   IOField "I/O field_37" at 183,323 size 90x29; Authorization "Commissioning"; FormatPattern 999; Unit  step
      ProcessValue <- "2110_BTCS_CNTRL_DB_BTCS_STEP"
   Button "HmiScreenItemData_10" at 43,323 size 137x29; TextOn 'Back'; TextOff 'BWTS Step'
   Button "HmiScreenItemData_51" at 43,358 size 137x29; TextOn 'Back'; TextOff 'BWTS State'
   Button "HmiScreenItemData_54" at 276,323 size 532x29; TextOn 'Back'; TextOff 'IGG STEP'; TextList "STEP LIST BTCS"
      ProcessValue <- "2110_BTCS_CNTRL_DB_BTCS_STEP"
   Button "HmiScreenItemData_55" at 276,358 size 532x29; TextOn 'Back'; TextOff 'IGG STEP'; TextList "STATE LIST BTCS"
      ProcessValue <- "2110_BTCS_CNTRL_DB_BTCS_STATE"
   Circle "Circle_2" at 421,496 size 26x26
      Appearance <- "80_From_HMI_BWT_BYPASS"
   Button "HmiScreenItemData_57" at 88,494 size 304x33; TextOn 'Back'; TextOff 'Ballast Water Treatment'; Authorization "Operate"
      on Press: InvertBit("80_From_HMI_BWT_BYPASS(1)"); ResetBit("80_From_HMI_CRG_BLNK_MODE(1)")
      Appearance <- "80_From_HMI_BWT_BYPASS(1)"
      ObjectEnable <- "100_GCU_AUTO_SEQ_DB_CRNT_STEP"
   Circle "Circle_3" at 421,534 size 26x26
      Appearance <- "80_From_HMI_CRG_BLNK_MODE"
   Button "HmiScreenItemData_58" at 88,532 size 304x33; TextOn 'Back'; TextOff 'Cargo Blanketing'; Authorization "Operate"
      on Press: InvertBit("80_From_HMI_CRG_BLNK_MODE(1)"); ResetBit("80_From_HMI_BWT_BYPASS(1)")
      Appearance <- "80_From_HMI_CRG_BLNK_MODE(1)"
      ObjectEnable <- "100_GCU_AUTO_SEQ_DB_CRNT_STEP"
   Button "HmiScreenItemData_56" at 41,461 size 425x27; TextOn 'Back'; TextOff 'Inert Gas Transfer Mode'
   Button "Button_7" at 817,526 size 79x32; TextOff '1'; Authorization "Operate"
      Appearance <- "504_Tank Grouping_DB2020_GROUP ACTIVE INT 1"
      on Press: function_b14e0dd5("504_Tank Grouping_DB2020_GROUP ACTIV 1", 0)
   Button "Button_8" at 817,560 size 79x32; TextOff '2'; Authorization "Operate"
      Appearance <- "504_Tank Grouping_DB2020_GROUP ACTIVE INT 2"
      on Press: function_b14e0dd5("504_Tank Grouping_DB2020_GROUP ACTIV 2", 0)
   Button "Button_9" at 493,539 size 100x23; TextOff 'TANK - 1P'; Authorization "Operate"
      on Press: function_b14e0dd5("504_Tank Grouping_DB2020_TANK ACTIV 2", 0)
      Appearance <- "504_Tank Grouping_DB2020_TANK ACTIV 2"
   Button "Button_14" at 493,571 size 100x23; TextOff 'TANK - 2P'; Authorization "Operate"
      on Press: function_b14e0dd5("504_Tank Grouping_DB2020_TANK ACTIV 4", 0)
      Appearance <- "504_Tank Grouping_DB2020_TANK ACTIV 4"
   Button "Button_15" at 493,603 size 100x23; TextOff 'TANK - 3P'; Authorization "Operate"
      on Press: function_b14e0dd5("504_Tank Grouping_DB2020_TANK ACTIV 6", 0)
      Appearance <- "504_Tank Grouping_DB2020_TANK ACTIV 6"
   Button "Button_16" at 493,636 size 100x23; TextOff 'TANK - 4P'; Authorization "Operate"
      on Press: function_b14e0dd5("504_Tank Grouping_DB2020_TANK ACTIV 8", 0)
      Appearance <- "504_Tank Grouping_DB2020_TANK ACTIV 8"
   Button "Button_17" at 493,668 size 100x23; TextOff 'TANK - 5P'; Authorization "Operate"
      on Press: function_b14e0dd5("504_Tank Grouping_DB2020_TANK ACTIV 10", 0)
      Appearance <- "504_Tank Grouping_DB2020_TANK ACTIV 10"
   Button "Button_18" at 493,700 size 100x23; TextOff 'TANK - 6P'; Authorization "Operate"
      on Press: function_b14e0dd5("504_Tank Grouping_DB2020_TANK ACTIV 12", 0)
      Appearance <- "504_Tank Grouping_DB2020_TANK ACTIV 12"
   Button "Button_19" at 493,733 size 100x23; TextOff 'TANK - APT'; Authorization "Operate"
      on Press: function_b14e0dd5("504_Tank Grouping_DB2020_TANK ACTIV 14", 0)
      Appearance <- "504_Tank Grouping_DB2020_TANK ACTIV 14"
   Button "Button_20" at 706,539 size 100x23; TextOff 'TANK - 1S'; Authorization "Operate"
      on Press: function_b14e0dd5("504_Tank Grouping_DB2020_TANK ACTIV 3", 0)
      Appearance <- "504_Tank Grouping_DB2020_TANK ACTIV 3"
   Button "Button_21" at 706,571 size 100x23; TextOff 'TANK - 2S'; Authorization "Operate"
      on Press: function_b14e0dd5("504_Tank Grouping_DB2020_TANK ACTIV 5", 0)
      Appearance <- "504_Tank Grouping_DB2020_TANK ACTIV 5"
   Button "Button_22" at 706,603 size 100x23; TextOff 'TANK - 3S'; Authorization "Operate"
      on Press: function_b14e0dd5("504_Tank Grouping_DB2020_TANK ACTIV 7", 0)
      Appearance <- "504_Tank Grouping_DB2020_TANK ACTIV 7"
   Button "Button_23" at 706,635 size 100x23; TextOff 'TANK - 4S'; Authorization "Operate"
      on Press: function_b14e0dd5("504_Tank Grouping_DB2020_TANK ACTIV 9", 0)
      Appearance <- "504_Tank Grouping_DB2020_TANK ACTIV 9"
   Button "Button_24" at 706,667 size 100x23; TextOff 'TANK - 5S'; Authorization "Operate"
      on Press: function_b14e0dd5("504_Tank Grouping_DB2020_TANK ACTIV 11", 0)
      Appearance <- "504_Tank Grouping_DB2020_TANK ACTIV 11"
   Button "Button_25" at 706,700 size 100x23; TextOff 'TANK - 6S'; Authorization "Operate"
      on Press: function_b14e0dd5("504_Tank Grouping_DB2020_TANK ACTIV 13", 0)
      Appearance <- "504_Tank Grouping_DB2020_TANK ACTIV 13"
   IOField "I/O field_38" at 183,358 size 90x29; Authorization "Commissioning"; FormatPattern 9; Unit  state
      ProcessValue <- "2110_BTCS_CNTRL_DB_BTCS_STATE"
   Switch "Switch_8" at 776,732 size 32x29; CaptionText 'Switch'; TextOn 'ON'; TextOff 'OFF'; Authorization "User administration"; PictureOff "Design_5_PilotLight_Green_Off"; PictureOn "Design_5_PilotLight_Green_On"
      on Change: InvertBit("80_From_HMI_Test Tank Request")
      ProcessValue <- "504_Tank Grouping_DB2020_RUN"
   Circle "Circle_31" at 621,507 size 20x20
      Appearance <- "504_Tank Grouping_DB2020_RUN TANK 1"
      Visibility <- "504_Tank Grouping_DB2020_RUN TANK 1"
   Circle "Circle_4" at 600,573 size 20x20
      Appearance <- "504_Tank Grouping_DB2020_GROUP of TANK 4"
   Circle "Circle_6" at 599,604 size 20x20
      Appearance <- "504_Tank Grouping_DB2020_GROUP of TANK 6"
   Circle "Circle_7" at 599,541 size 20x20
      Appearance <- "504_Tank Grouping_DB2020_GROUP of TANK 2"
   Circle "Circle_8" at 599,669 size 20x20
      Appearance <- "504_Tank Grouping_DB2020_GROUP of TANK 10"
   Circle "Circle_10" at 599,637 size 20x20
      Appearance <- "504_Tank Grouping_DB2020_GROUP of TANK 8"
   Circle "Circle_11" at 599,734 size 20x20
      Appearance <- "504_Tank Grouping_DB2020_GROUP of TANK 14"
   Circle "Circle_12" at 599,701 size 20x20
      Appearance <- "504_Tank Grouping_DB2020_GROUP of TANK 12"
   IOField "I/O field_8" at 599,544 size 20x14; FormatPattern 99
      ProcessValue <- "504_Tank Grouping_DB2020_GROUP of TANK 2"
   IOField "I/O field_9" at 599,576 size 20x14; FormatPattern 99
      ProcessValue <- "504_Tank Grouping_DB2020_GROUP of TANK 4"
   IOField "I/O field_26" at 599,607 size 20x14; FormatPattern 99
      ProcessValue <- "504_Tank Grouping_DB2020_GROUP of TANK 6"
   IOField "I/O field_28" at 599,640 size 20x14; FormatPattern 99
      ProcessValue <- "504_Tank Grouping_DB2020_GROUP of TANK 8"
   IOField "I/O field_30" at 599,672 size 20x14; FormatPattern 99
      ProcessValue <- "504_Tank Grouping_DB2020_GROUP of TANK 10"
   IOField "I/O field_33" at 599,704 size 20x14; FormatPattern 99
      ProcessValue <- "504_Tank Grouping_DB2020_GROUP of TANK 12"
   IOField "I/O field_35" at 599,737 size 20x14; FormatPattern 99
      ProcessValue <- "504_Tank Grouping_DB2020_GROUP of TANK 14"
   Circle "Circle_13" at 678,573 size 20x20
      Appearance <- "504_Tank Grouping_DB2020_GROUP of TANK 5"
   Circle "Circle_14" at 678,603 size 20x20
      Appearance <- "504_Tank Grouping_DB2020_GROUP of TANK 7"
   Circle "Circle_15" at 678,541 size 20x20
      Appearance <- "504_Tank Grouping_DB2020_GROUP of TANK 3"
   Circle "Circle_16" at 678,668 size 20x20
      Appearance <- "504_Tank Grouping_DB2020_GROUP of TANK 11"
   Circle "Circle_17" at 678,636 size 20x20
      Appearance <- "504_Tank Grouping_DB2020_GROUP of TANK 9"
   Circle "Circle_18" at 678,701 size 20x20
      Appearance <- "504_Tank Grouping_DB2020_GROUP of TANK 13"
   IOField "I/O field_23" at 678,544 size 20x14; FormatPattern 99
      ProcessValue <- "504_Tank Grouping_DB2020_GROUP of TANK 3"
   IOField "I/O field_24" at 678,576 size 20x14; FormatPattern 99
      ProcessValue <- "504_Tank Grouping_DB2020_GROUP of TANK 5"
   IOField "I/O field_27" at 678,606 size 20x14; FormatPattern 99
      ProcessValue <- "504_Tank Grouping_DB2020_GROUP of TANK 7"
   IOField "I/O field_29" at 678,639 size 20x14; FormatPattern 99
      ProcessValue <- "504_Tank Grouping_DB2020_GROUP of TANK 9"
   IOField "I/O field_32" at 678,671 size 20x14; FormatPattern 99
      ProcessValue <- "504_Tank Grouping_DB2020_GROUP of TANK 11"
   IOField "I/O field_34" at 678,704 size 20x14; FormatPattern 99
      ProcessValue <- "504_Tank Grouping_DB2020_GROUP of TANK 13"
   Circle "Circle_32" at 621,540 size 20x20
      Appearance <- "504_Tank Grouping_DB2020_RUN TANK 2"
      Visibility <- "504_Tank Grouping_DB2020_RUN TANK 2"
   Circle "Circle_33" at 656,540 size 20x20
      Appearance <- "504_Tank Grouping_DB2020_RUN TANK 3"
      Visibility <- "504_Tank Grouping_DB2020_RUN TANK 3"
   Circle "Circle_34" at 621,572 size 20x20
      Appearance <- "504_Tank Grouping_DB2020_RUN TANK 4"
      Visibility <- "504_Tank Grouping_DB2020_RUN TANK 4"
   Circle "Circle_35" at 656,572 size 20x20
      Appearance <- "504_Tank Grouping_DB2020_RUN TANK 5"
      Visibility <- "504_Tank Grouping_DB2020_RUN TANK 5"
   Circle "Circle_36" at 621,604 size 20x20
      Appearance <- "504_Tank Grouping_DB2020_RUN TANK 6"
      Visibility <- "504_Tank Grouping_DB2020_RUN TANK 6"
   Circle "Circle_37" at 656,604 size 20x20
      Appearance <- "504_Tank Grouping_DB2020_RUN TANK 7"
      Visibility <- "504_Tank Grouping_DB2020_RUN TANK 7"
   Circle "Circle_38" at 621,636 size 20x20
      Appearance <- "504_Tank Grouping_DB2020_RUN TANK 8"
      Visibility <- "504_Tank Grouping_DB2020_RUN TANK 8"
   Circle "Circle_39" at 656,636 size 20x20
      Appearance <- "504_Tank Grouping_DB2020_RUN TANK 9"
      Visibility <- "504_Tank Grouping_DB2020_RUN TANK 9"
   Circle "Circle_40" at 621,668 size 20x20
      Appearance <- "504_Tank Grouping_DB2020_RUN TANK 10"
      Visibility <- "504_Tank Grouping_DB2020_RUN TANK 10"
   Circle "Circle_41" at 656,668 size 20x20
      Appearance <- "504_Tank Grouping_DB2020_RUN TANK 11"
      Visibility <- "504_Tank Grouping_DB2020_RUN TANK 11"
   Circle "Circle_42" at 621,701 size 20x20
      Appearance <- "504_Tank Grouping_DB2020_RUN TANK 12"
      Visibility <- "504_Tank Grouping_DB2020_RUN TANK 12"
   Circle "Circle_43" at 656,701 size 20x20
      Appearance <- "504_Tank Grouping_DB2020_RUN TANK 13"
      Visibility <- "504_Tank Grouping_DB2020_RUN TANK 13"
   Circle "Circle_44" at 621,733 size 20x20
      Appearance <- "504_Tank Grouping_DB2020_RUN TANK 14"
      Visibility <- "504_Tank Grouping_DB2020_RUN TANK 14"
   TextField "Text field_7" at 648,740 size 136x18; Text 'Test Tank Request'
   Rectangle "Rectangle_6" at 816,488 size 82x37
      Visibility <- "504_Tank Grouping_DB2020_SetGroupSR"
   Button "Button_13" at 819,491 size 76x31; TextOff 'Set Group'; Authorization "Parameter Change"
      Appearance <- "504_Tank Grouping_DB2020_GROUP SET"
      on Press: function_b14e0dd5("504_Tank Grouping_DB2020_SetGroup", 0)
   Button "HmiScreenItemData_5" at 41,576 size 426x27; TextOn 'Back'; TextOff 'Automatic Gas to Tank Valves Cycling'
   Button "HmiScreenItemData_19" at 371,722 size 83x35; TextOn 'ENABLE'; TextOff 'Enable'; Authorization "Operating Mode"
      on Press: InvertBit("504_Tank Grouping_DB2020_Valve Cycle_Enable")
      Appearance <- "504_Tank Grouping_DB2020_Valve Cycle_Enable"
   TextField "Text field_8" at 54,652 size 254x18; Text 'Gas to Tank Valves Cycle Frequency'
   TextField "Text field_9" at 54,690 size 233x18; Text 'Gas to Tank Valves Cycle Length'
   TextField "Text field_10" at 54,618 size 85x18; Text 'Description'
   TextField "Text field_12" at 311,618 size 67x18; Text 'Setpoint'
   IOField "I/O field_39" at 310,649 size 70x28; Authorization "Operate"; FormatPattern 999; Unit h
      ProcessValue <- "504_Tank Grouping_DB2020_Valve Cycle_Period"
   IOField "I/O field_40" at 310,685 size 70x28; Authorization "Operate"; FormatPattern 9999; Unit s
      ProcessValue <- "504_Tank Grouping_DB2020_Valve Cycle_Length"
   TextField "Text field_13" at 385,618 size 58x18; Text 'Elapsed'
   IOField "I/O field_41" at 384,649 size 70x28; Authorization "Operate"; FormatPattern 999; Unit h
      ProcessValue <- "504_Tank Grouping_DB2020_Cycle Period_ET"
   IOField "I/O field_42" at 384,685 size 70x28; Authorization "Operate"; FormatPattern 9999; Unit s
      ProcessValue <- "504_Tank Grouping_DB2020_Cycle Length_ET"
   IOField "I/O field_48" at 1172,169 size 33x28; Authorization "User administration"; FormatPattern 99; Unit h
      ProcessValue <- "Sequence Times_DB_Treatment Timer_Hours Left"
   IOField "I/O field_51" at 1140,169 size 33x28; Authorization "User administration"; FormatPattern 99; Unit d
      ProcessValue <- "Sequence Times_DB_Treatment Timer_Days Left"
   IOField "I/O field_52" at 1204,169 size 35x28; Authorization "User administration"; FormatPattern 99; Unit m
      ProcessValue <- "Sequence Times_DB_Treatment Timer_Minutes Left"
   IOField "I/O field_43" at 1156,201 size 83x28; Authorization "User administration"; FormatPattern 999; Unit  min
      ProcessValue <- "504_Tank Grouping_DB2020_Diff Time Remain"
      Visibility <- "AlwaysTRUE"
   IOField "I/O field_44" at 1204,233 size 35x28; Authorization "User administration"; FormatPattern 99; Unit m
      ProcessValue <- "Sequence Times_DB_Pre-Dwell Timer_Minutes Left"
   IOField "I/O field_45" at 1172,233 size 33x28; Authorization "User administration"; FormatPattern 99; Unit h
      ProcessValue <- "Sequence Times_DB_Pre-Dwell Timer_Hours Left"
   IOField "I/O field_46" at 1140,233 size 33x28; Authorization "User administration"; FormatPattern 99; Unit d
      ProcessValue <- "Sequence Times_DB_Pre-Dwell Timer_Days Left"
   IOField "I/O field_47" at 1040,132 size 92x28; Authorization "Operating Mode"; FormatPattern 999.9; Unit  Days
      ProcessValue <- "Sequence Times_DB_Jurney Time"
   IOField "I/O field_49" at 1072,169 size 33x28; Authorization "User administration"; FormatPattern 99; Unit h
      ProcessValue <- "Sequence Times_DB_Treatment Timer_Hours"
   IOField "I/O field_50" at 1040,169 size 33x28; Authorization "User administration"; FormatPattern 99; Unit d
      ProcessValue <- "Sequence Times_DB_Treatment Timer_Days"
   IOField "I/O field_53" at 1104,169 size 35x28; Authorization "User administration"; FormatPattern 99; Unit m
      ProcessValue <- "Sequence Times_DB_Treatment Timer_Minutes"
   IOField "I/O field_54" at 1172,132 size 33x28; Authorization "User administration"; FormatPattern 99; Unit h
      ProcessValue <- "Sequence Times_DB_Jurney Timer_Hours Left"
   IOField "I/O field_55" at 1133,132 size 40x28; Authorization "User administration"; FormatPattern 999; Unit d
      ProcessValue <- "Sequence Times_DB_Jurney Timer_Days Left"
   IOField "I/O field_56" at 1204,132 size 35x28; Authorization "User administration"; FormatPattern 99; Unit m
      ProcessValue <- "Sequence Times_DB_Jurney Timer_Minutes Left"
   IOField "I/O field_57" at 1040,233 size 79x28; Authorization "Commissioning"; FormatPattern 9999.9; Unit  Hrs
      ProcessValue <- "Sequence Times_DB_Pre-Dwell Time"
   IOField "I/O field_58" at 1040,267 size 79x28; Authorization "Commissioning"; FormatPattern 999.9; Unit  Hrs
      ProcessValue <- "Sequence Times_DB_De-Ox Time"
   IOField "I/O field_59" at 1204,267 size 35x28; Authorization "User administration"; FormatPattern 99; Unit m
      ProcessValue <- "Sequence Times_DB_De-Ox Timer_Minutes Left"
   IOField "I/O field_60" at 1172,267 size 33x28; Authorization "User administration"; FormatPattern 99; Unit h
      ProcessValue <- "Sequence Times_DB_De-Ox Timer_Hours Left"
   IOField "I/O field_61" at 1140,267 size 33x28; Authorization "User administration"; FormatPattern 99; Unit d
      ProcessValue <- "Sequence Times_DB_De-Ox Timer_Days Left"
   IOField "I/O field_62" at 1040,301 size 79x28; Authorization "Commissioning"; FormatPattern 999.9; Unit  Hrs
      ProcessValue <- "Sequence Times_DB_De-Ox SP Time"
   IOField "I/O field_63" at 1040,335 size 79x28; Authorization "Commissioning"; FormatPattern 999.9; Unit  Hrs
      ProcessValue <- "Sequence Times_DB_Dwell Time"
   IOField "I/O field_64" at 1204,335 size 35x28; Authorization "User administration"; FormatPattern 99; Unit m
      ProcessValue <- "Sequence Times_DB_Dwell Timer_Minutes Left"
   IOField "I/O field_65" at 1172,335 size 33x28; Authorization "User administration"; FormatPattern 99; Unit h
      ProcessValue <- "Sequence Times_DB_Dwell Timer_Hours Left"
   IOField "I/O field_66" at 1140,335 size 33x28; Authorization "User administration"; FormatPattern 99; Unit d
      ProcessValue <- "Sequence Times_DB_Dwell Timer_Days Left"
   IOField "I/O field_2" at 1040,369 size 79x28; Authorization "Commissioning"; FormatPattern 999.9; Unit  Hrs
      ProcessValue <- "Sequence Times_DB_Re-Ox Time"
   IOField "I/O field_67" at 1204,369 size 35x28; Authorization "User administration"; FormatPattern 99; Unit m
      ProcessValue <- "Sequence Times_DB_Re-Ox Timer_Minutes Left"
   IOField "I/O field_68" at 1172,369 size 33x28; Authorization "User administration"; FormatPattern 99; Unit h
      ProcessValue <- "Sequence Times_DB_Re-Ox Timer_Hours Left"
   IOField "I/O field_69" at 1140,369 size 33x28; Authorization "User administration"; FormatPattern 99; Unit d
      ProcessValue <- "Sequence Times_DB_Re-Ox Timer_Days Left"
   IOField "I/O field_70" at 1040,403 size 79x28; Authorization "Commissioning"; FormatPattern 999.9; Unit  Hrs
      ProcessValue <- "Sequence Times_DB_Post-Dwell Time"
   IOField "I/O field_71" at 1204,403 size 35x28; Authorization "User administration"; FormatPattern 99; Unit m
      ProcessValue <- "Sequence Times_DB_Post-Dwell Timer_Minutes Left"
   IOField "I/O field_72" at 1172,403 size 33x28; Authorization "User administration"; FormatPattern 99; Unit h
      ProcessValue <- "Sequence Times_DB_Post-Dwell Timer_Hours Left"
   IOField "I/O field_73" at 1140,403 size 33x28; Authorization "User administration"; FormatPattern 99; Unit d
      ProcessValue <- "Sequence Times_DB_Post-Dwell Timer_Days Left"
   TextField "Text field_15" at 621,419 size 156x18; Text 'Treatment Timer Test'
      Visibility <- "user_group"
   Circle "Circle_5" at 599,507 size 20x20
      Appearance <- "504_Tank Grouping_DB2020_GROUP of TANK 1"
   IOField "I/O field_7" at 599,510 size 20x14; FormatPattern 99
      ProcessValue <- "504_Tank Grouping_DB2020_GROUP of TANK 1"
   Button "HmiScreenItemData_50" at 1156,297 size 83x35; TextOn 'Back'; TextOff 'Boost'; Authorization "Commissioning"
      on Press: InvertBit("Sequence Times_DB_Boost")
      Visibility <- "user_group"
      Appearance <- "Sequence Times_DB_Boost"
   TextField "Text field_16" at 38,419 size 76x18; Text 'HeartBeat'
      Visibility <- "user_group"
   TextField "Text field_18" at 201,422 size 107x18; Text 'PLC HeartBeat'
      Visibility <- "user_group"
   Circle "Circle_45" at 6,412 size 26x26
      Appearance <- "IGG HMI HEART BEAT"
   Circle "Circle_46" at 166,414 size 26x26
      Appearance <- "IGG PLC HEART BEAT"
   Switch "Switch_1" at 774,411 size 32x29; CaptionText 'Switch'; TextOn 'ON'; TextOff 'OFF'; Authorization "User administration"; PictureOff "Design_5_PilotLight_Green_Off"; PictureOn "Design_5_PilotLight_Green_On"
      on Change: InvertBit("80_From_HMI_Jurney Start Simulator")
      Visibility <- "user_group"
      ProcessValue <- "80_From_HMI_Jurney Start Simulator"
   TextField "Text field_19" at 445,403 size 133x18; Text 'Log IGG Simulator'
      Visibility <- "user_group"
   Switch "Switch_2" at 568,393 size 32x29; CaptionText 'Switch'; TextOn 'ON'; TextOff 'OFF'; Authorization "User administration"; PictureOff "Design_5_PilotLight_Green_Off"; PictureOn "Design_5_PilotLight_Green_On"
      on Change: InvertBit("68_Sys_Status_Data_LOG IGG Simulator")
      Visibility <- "user_group"
      ProcessValue <- "68_Sys_Status_Data_LOG IGG Simulator"
   TextField "Text field_20" at 445,435 size 136x18; Text 'Log GCU Simulator'
      Visibility <- "user_group"
   Switch "Switch_3" at 568,425 size 32x29; CaptionText 'Switch'; TextOn 'ON'; TextOff 'OFF'; Authorization "User administration"; PictureOff "Design_5_PilotLight_Green_Off"; PictureOn "Design_5_PilotLight_Green_On"
      on Change: InvertBit("68_Sys_Status_Data_LOG GCU Simulator")
      Visibility <- "user_group"
      ProcessValue <- "68_Sys_Status_Data_LOG GCU Simulator"
   Button "Button_5" at 53,722 size 210x35; TextOff 'PGC Setpoint Protection'
      on Press: function_efd93a16("PGC Setpoint Protection", 400, 200, -1, -1, 1)
   Button "Button_26" at 280,114 size 209x107; TextOff 'Text'
      on Release: function_efd93a16("Salinity - Acceptance", 168, 315, -1, 0, 1)
      Visibility <- "2068_Sys_Status_Data_SAL_VALID"
   Button "Button_27" at 283,115 size 204x107; TextOff 'Text'
      on Release: function_efd93a16("Tank Times", 300, 200, -1, 0, 1)
      Visibility <- "2068_Sys_Status_Data_Times Visibil"
   Group "Group_1" at 909,732 size 329x37
   IOField "I/O field_74" at 1172,201 size 33x28; Authorization "User administration"; FormatPattern 99; Unit h
      ProcessValue <- "Sequence Times_DB_Offset Timer_Hours Left"
   IOField "I/O field_75" at 1140,201 size 33x28; Authorization "User administration"; FormatPattern 99; Unit d
      ProcessValue <- "Sequence Times_DB_Offset Timer_Days Left"
   IOField "I/O field_76" at 1204,201 size 35x28; Authorization "User administration"; FormatPattern 99; Unit m
      ProcessValue <- "Sequence Times_DB_Offset Timer_Minutes Left"
   Circle "Circle_23" at 762,90 size 24x24
      Appearance <- "2110_BTCS_CNTRL_DB_BTCS_STEP"
   Circle "Circle_24" at 762,119 size 24x24
      Appearance <- "100_GCU_AUTO_SEQ_DB_CRNT_STEP"
   Circle "Circle_25" at 762,149 size 24x24
      Appearance <- "2110_BTCS_CNTRL_DB_BTCS_STEP"
   Circle "Circle_26" at 762,179 size 24x24
      Appearance <- "2110_BTCS_CNTRL_DB_BTCS_STEP"
   Circle "Circle_27" at 762,209 size 24x24
      Appearance <- "100_GCU_AUTO_SEQ_DB_CRNT_STEP"
   Circle "Circle_28" at 762,239 size 24x24
      Appearance <- "2110_BTCS_CNTRL_DB_BTCS_STEP"
   Circle "Circle_29" at 762,269 size 24x24
      Appearance <- "2110_BTCS_CNTRL_DB_BTCS_STEP"
   TextField "Text field_34" at 980,733 size 187x35; Text 'TIMES VALID'
      Visibility <- "2102_TIME_CALCS_DB_TIMES_VALID"
   TextField "Text field_4" at 909,732 size 329x37; Text 'TIMES INVALID'
      Visibility <- "2102_TIME_CALCS_DB_TIMES_VALID"
   Rectangle "Rectangle_27" at 921,659 size 322x40
      Visibility <- "2068_Sys_Status_Data_SAL_CNF_CHK"
   TextField "Text field_62" at 925,664 size 156x30; Text 'Confirm Salinity? :'
      Visibility <- "2068_Sys_Status_Data_SAL_CNF_CHK"
   Button "Button_6" at 1086,664 size 67x30; TextOff 'YES'
      on Press: function_b14e0dd5("80_From_HMI_LOW_SAL_ACPT", 0)
      Visibility <- "2068_Sys_Status_Data_SAL_CNF_CHK"
   Button "Button_3" at 1166,664 size 67x30; TextOff 'NO'
      on Press: function_b14e0dd5("80_From_HMI_LOW_SAL_RJCT", 0)
      Visibility <- "2068_Sys_Status_Data_SAL_CNF_CHK"
   Rectangle "Rectangle_28" at 916,659 size 327x40
      Visibility <- "2100_AUTO_SEQ_DB_SEQ_RNG"
      Appearance <- "2102_TIME_CALCS_DB_RE_OX_SP_TMR_DN"
   TextField "Text field_49" at 920,664 size 211x30; Text 'Salinity Value :'
      Visibility <- "2100_AUTO_SEQ_DB_SEQ_RNG"
   IOField "I/O field_36" at 1131,664 size 95x30; Authorization "Operate"; FormatPattern 99.9; Unit psu
      Visibility <- "2100_AUTO_SEQ_DB_SEQ_RNG"
      ProcessValue <- "80_From_HMI_SAL_VALUE"

PopupScreen "SD Card overflow" 665x230
   Button "Button_1" at 0,0 size 665x230; TextOff 'Data Logging SD Card Memory Full'
      on Click: function_efd93a16("SD Card overflow", 0, 0, -1, -1, 1)
      on Press: ResetBit("Logging SD Card Overflow")

PopupScreen "Salinity - Fresh Water Alert" 1280x800
   Button "Button_1" at 115,225 size 1050x284; TextOff 'NOTE: BALLAST WATER SALINITY IS FRESH WATER LEVEL This System Is Not Certified For FRESH WATER Treatment. Do Wish To Continue Ballast Water Treatment?'
   Button "Button_2" at 666,514 size 105x50; TextOff 'NO'
      on Release: ActivateScreen("Balast Water Treatment Setup", 0)
      on Press: function_b14e0dd5("80_From_HMI_LOW_SAL_RJCT", 0)
   Button "Button_3" at 500,514 size 105x50; TextOff 'YES'
      on Release: ActivateScreen("Balast Water Treatment Setup", 0)
      on Press: function_b14e0dd5("80_From_HMI_LOW_SAL_ACPT", 0)

screen "Main Page" 1280x800, template "Template"
   GraphicView "Graphic view_49" at 158,415 size 30x45; Picture "Graphic_72"
   GraphicView "Graphic view_20" at 140,368 size 380x356; Picture "IGG_6"
   GraphicView "Graphic view_62" at 134,449 size 92x8; Picture "Graphic_20"
   GraphicView "Graphic view_5" at 464,423 size 90x19; Picture "Graphic_82"
   GraphicView "Graphic view_41" at 228,459 size 9x40; Picture "Graphic_57"
   GraphicView "Graphic view_40" at 222,449 size 15x13; Picture "Graphic_41"
   GraphicView "Graphic view_21" at 210,503 size 17x7; Picture "Graphic_63"
   GraphicView "Graphic view_22" at 207,499 size 8x9; Picture "Graphic_64"
   GraphicView "Graphic view_23" at 206,399 size 6x104; Picture "Graphic_70"
   GraphicView "Graphic view_39" at 138,535 size 6x7; Picture "Graphic_70"
   GraphicView "Graphic view_38" at 139,539 size 7x9; Picture "Graphic_64"
   GraphicView "Graphic view_18" at 204,397 size 9x10; Picture "Graphic_67"
   Group "Group_3" at 158,415 size 30x41; Picture "Graphic_72"
   GraphicView "Graphic view_65" at 144,542 size 8x6; Picture "Graphic_63"
   GraphicView "Graphic view_69" at 295,453 size 14x15; Picture "Graphic_36"
   GraphicView "Graphic view_70" at 335,462 size 14x15; Picture "Graphic_36"
   GraphicView "Graphic view_71" at 251,443 size 14x17; Picture "Graphic_79"
   GraphicView "Graphic view_36" at 517,373 size 35x50; Picture "Graphic_108"
   GraphicView "Graphic view_4" at 333,376 size 31x49; Picture "Graphic_108"
   GraphicView "Graphic view_72" at 387,407 size 14x17; Picture "Graphic_36"
   GraphicView "Graphic view_37" at 136,525 size 8x11; Picture "Graphic_67"
   GraphicView "Graphic view_89" at 440,407 size 14x17; Picture "Graphic_36"
   Line "Line_4" at 226,517 size 2x15
      Visibility <- "14_DQ_Data_X001ControlOut"
   GraphicView "Graphic view_84" at 215,511 size 27x55; Picture "Graphic_129"
      Visibility <- "102_Pilot_Burner_DB_FLM_DET"
   GraphicView "Graphic view_90" at 488,409 size 14x15; Picture "Graphic_36"
   GraphicView "Graphic view_1" at 342,415 size 18x41; Picture "Graphic_17"
   GraphicView "Graphic view_60" at 526,412 size 18x41; Picture "Graphic_17"
   GraphicView "Graphic view_82" at 210,499 size 167x147; Picture "Graphic_130"
      Visibility <- "103_Main_Burner_DB_DN_OK(1)"
   IOField "I/O field_17" at 231,558 size 46x17; FormatPattern 999; Unit %
      Visibility <- "10 DI_DATA_FD001_OK"
      ProcessValue <- "12_AI_Data_FD001FlameSignalIn"
   GraphicView "Graphic view_63" at 133,396 size 75x7; Picture "Graphic_63"
   GraphicView "Graphic view_25" at 659,340 size 25x46; Picture "Graphic_148"
   Group "Group_10" at 659,340 size 26x47; Picture "Graphic_148"
   Group "Group_11" at 649,372 size 56x37; Picture "Graphic_224"
   GraphicView "Graphic view_26" at 649,373 size 55x36; Picture "Graphic_224"
   GraphicView "Graphic view_27" at 569,502 size 205x15; Picture "Graphic_232"
   GraphicView "Graphic view_3" at 78,471 size 64x14; Picture "Graphic_82"
   GraphicView "Graphic view_19" at 776,616 size 64x10; Picture "Graphic_82"
   GraphicIOField "Graphic I/O field_2" at 0,485 size 128x131; PictureList "IA Compressor_1"
      ProcessValue <- "82_To_HMI_CA Blower Animation"
   GraphicView "Graphic view_7" at 700,602 size 119x212; Picture "Graphic_150"
   Group "Group" at 133,368 size 421x356; Picture "Graphic_20"
   GraphicView "Graphic view_2" at 821,493 size 449x266; Picture "Graphic_185"
   GraphicView "Graphic view_6" at 68,470 size 18x21; Picture "Graphic_66"
   GraphicView "Graphic view_8" at 41,328 size 96x93; Picture "Graphic_246"
   GraphicView "Graphic view_14" at 630,544 size 17x40; Picture "Graphic_271"
   GraphicView "Graphic view_15" at 570,390 size 205x15; Picture "Graphic_232"
   GraphicView "Graphic view_16" at 561,391 size 26x27; Picture "Graphic_178"
   GraphicView "Graphic view_17" at 757,380 size 17x35; Picture "Graphic_280"
   GraphicView "Graphic view_9" at 525,539 size 156x153; Picture "Graphic_251"
   GraphicView "Graphic view_24" at 561,407 size 14x167; Picture "Graphic_231"
   GraphicView "Graphic view_11" at 555,635 size 21x22; Picture "Graphic_265"
   GraphicView "Graphic view_12" at 555,653 size 29x31; Picture "Graphic_266"
   GraphicView "Graphic view_13" at 572,667 size 133x18; Picture "Graphic_232"
   GraphicView "Graphic view_10" at 549,422 size 26x38; Picture "Graphic_169"
   Group "Group_12" at 649,340 size 56x69; Picture "Graphic_148"
   GraphicView "Graphic view_28" at 756,492 size 17x35; Picture "Graphic_280"
   Group "Group_4" at 648,452 size 56x69; Picture "Graphic_148"
   GraphicView "Graphic view_29" at 658,452 size 25x46; Picture "Graphic_148"
   Group "Group_1" at 658,452 size 26x47; Picture "Graphic_148"
   Group "Group_2" at 648,484 size 56x37; Picture "Graphic_224"
   GraphicView "Graphic view_30" at 648,485 size 55x36; Picture "Graphic_224"

screen "GCU Analogue Inputs" 1280x800, template "Template"
   on GenerateScreen: "TitleUpdater"()
   Button "HmiScreenItemData_1" at 1,1 size 150x43; TextOn 'Back'; TextOff 'Commissioning'
      on Release: ActivateScreen("Commissioning Main Page", 0)
   TextField "Text field_6" at 7,150 size 53x22; Text 'IW800'
   TextField "Text field_8" at 7,270 size 53x22; Text 'IW806'
   TextField "Text field_10" at 7,310 size 53x22; Text 'IW808'
   TextField "Text field_12" at 7,430 size 53x22; Text 'IW814'
   TextField "Text field_30" at 1203,124 size 74x20; Text 'High High'
   TextField "Text field_54" at 649,719 size 228x62; Text 'Note: CSW = Cooling Sea Water'
   TextField "Text field_32" at 7,231 size 53x22; Text 'IW804'
   TextField "Text field_34" at 7,391 size 53x22; Text 'IW812'
   TextField "Text field_36" at 8,191 size 53x22; Text 'IW802'
   TextField "Text field_38" at 8,349 size 53x22; Text 'IW810'
   AlarmView "Alarm view_1" at 0,777 size 1280x23
   IOField "I/O field_62" at 1208,191 size 60x22; FormatPattern 9.9
      ProcessValue <- "84_Setpoints_E400_PT002_HighHigh"
   IOField "I/O field_61" at 1140,191 size 60x22; FormatPattern 9.9
      ProcessValue <- "84_Setpoints_E400_PT002_High"
   TextField "Text field_82" at 60,150 size 220x22; Text 'LIT304 GCU LEVEL'
   TextField "Text field_90" at 286,124 size 64x20; Text 'Reading'
   IOField "I/O field_2" at 287,150 size 70x22; FormatPattern 999; Unit  %
      ProcessValue <- "12_AI_Data_LIT_304_SCALED"
   TextField "Text field_1" at 359,124 size 68x20; Text 'Low Low'
   IOField "I/O field_1" at 361,150 size 60x22; Authorization "Parameter Change"; FormatPattern 999
      ProcessValue <- "19_AUTO_CMNDS_Data_LIT304_CMND_LowLow"
   TextField "Text field_2" at 442,124 size 37x20; Text 'Low'
   IOField "I/O field_3" at 429,150 size 60x22; Authorization "Parameter Change"; FormatPattern 999
      ProcessValue <- "19_AUTO_CMNDS_Data_LIT304_CMND_Low"
   TextField "Text field_3" at 509,124 size 37x20; Text 'High'
   IOField "I/O field_4" at 497,150 size 60x22; Authorization "Parameter Change"; FormatPattern 999
      ProcessValue <- "19_AUTO_CMNDS_Data_LIT304_CMND_High"
   TextField "Text field_4" at 561,124 size 74x20; Text 'High High'
   IOField "I/O field_5" at 565,150 size 60x22; Authorization "Parameter Change"; FormatPattern 999
      ProcessValue <- "19_AUTO_CMNDS_Data_LIT304_CMND_HighHigh"
   TextField "Text field_5" at 434,100 size 76x20; Text 'Setpoints'
   TextField "Text field_7" at 60,270 size 220x22; Text 'TIT406 GAS TO DECK TEMP'
   IOField "I/O field_6" at 287,270 size 70x22; FormatPattern s999; Unit  °C
      ProcessValue <- "12_AI_Data_TIT_406_SCALED"
   IOField "I/O field_7" at 361,270 size 60x22; FormatPattern 999
   IOField "I/O field_8" at 429,270 size 60x22; FormatPattern 999
   IOField "I/O field_9" at 497,270 size 60x22; Authorization "Parameter Change"; FormatPattern 999
      ProcessValue <- "84_Setpoints_TIT406_High"
   IOField "I/O field_10" at 565,270 size 60x22; Authorization "Parameter Change"; FormatPattern 999
      ProcessValue <- "84_Setpoints_TIT406_HighHigh"
   TextField "Text field_9" at 60,310 size 220x22; Text 'CV405 POSITION'
   IOField "I/O field_11" at 287,310 size 70x22; FormatPattern 999; Unit  %
      ProcessValue <- "12_AI_Data_CV_405_SCALED"
   IOField "I/O field_12" at 361,310 size 60x22; Authorization "Parameter Change"; FormatPattern 999
   IOField "I/O field_13" at 429,310 size 60x22; Authorization "Parameter Change"; FormatPattern 999
   IOField "I/O field_14" at 497,310 size 60x22; Authorization "Parameter Change"; FormatPattern 999
   IOField "I/O field_15" at 565,310 size 60x22; Authorization "Parameter Change"; FormatPattern 999
   TextField "Text field_11" at 60,430 size 220x22; Text 'PIT348 GCU CSW PRESS'
   IOField "I/O field_16" at 287,430 size 70x22; FormatPattern s9.9; Unit  Barg
      ProcessValue <- "12_AI_Data_PIT_348_SCALED"
   IOField "I/O field_17" at 361,430 size 60x22; FormatPattern 9.9
      ProcessValue <- "84_Setpoints_PIT348_LowLow"
   IOField "I/O field_18" at 429,430 size 60x22; FormatPattern 9.9
      ProcessValue <- "84_Setpoints_PIT348_Low"
   IOField "I/O field_19" at 497,430 size 60x22; FormatPattern 9.9
      ProcessValue <- "84_Setpoints_PIT348_High"
   IOField "I/O field_20" at 565,430 size 60x22; FormatPattern 9.9
      ProcessValue <- "84_Setpoints_PIT348_HighHigh"
   TextField "Text field_21" at 703,151 size 220x22; Text 'PIT353 RECIRC FCW PRESS'
   IOField "I/O field_41" at 930,151 size 70x22; FormatPattern s9.9; Unit  Barg
      ProcessValue <- "12_AI_Data_PIT_353_SCALED"
   IOField "I/O field_42" at 1004,151 size 60x22; Authorization "Commissioning"; FormatPattern 9.9
      ProcessValue <- "19_AUTO_CMNDS_Data_PIT353_CMND_LowLow"
   IOField "I/O field_43" at 1072,151 size 60x22; Authorization "Commissioning"; FormatPattern 9.9
      ProcessValue <- "19_AUTO_CMNDS_Data_PIT353_CMND_Low"
   IOField "I/O field_44" at 1140,151 size 60x22; FormatPattern 9.9
      ProcessValue <- "19_AUTO_CMNDS_Data_PIT353_CMND_High"
   IOField "I/O field_45" at 1208,151 size 60x22; FormatPattern 9.9
      ProcessValue <- "19_AUTO_CMNDS_Data_PIT353_CMND_HighHigh"
   TextField "Text field_22" at 650,151 size 53x22; Text 'IW816'
   TextField "Text field_23" at 703,191 size 220x22; Text 'E400 PT002 PGC PRESS'
   IOField "I/O field_46" at 930,191 size 70x22; FormatPattern s9.9; Unit  Barg
      ProcessValue <- "12_AI_Data_E_400_PT002_SCALED"
   TextField "Text field_24" at 650,191 size 53x22; Text 'IW818'
   TextField "Text field_26" at 928,124 size 64x20; Text 'Reading'
   TextField "Text field_27" at 1001,124 size 68x20; Text 'Low Low'
   TextField "Text field_28" at 1082,124 size 37x20; Text 'Low'
   TextField "Text field_29" at 1150,124 size 37x20; Text 'High'
   TextField "Text field_31" at 1076,100 size 76x20; Text 'Setpoints'
   TextField "Text field_51" at 703,231 size 220x22; Text 'E400 TT002 PGC TEMP'
   IOField "I/O field_101" at 930,231 size 70x22; FormatPattern s999; Unit  °C
      ProcessValue <- "12_AI_Data_E_400_TE002_SCALED"
   TextField "Text field_56" at 650,231 size 53x22; Text 'IW820'
   TextField "Text field_57" at 703,271 size 220x22; Text 'SL400 BALLAST SALINITY'
   IOField "I/O field_106" at 930,271 size 70x22; FormatPattern 999; Unit  %
      ProcessValue <- "12_AI_Data_SL_400_SCALED"
   IOField "I/O field_107" at 1004,271 size 60x22; FormatPattern 999
   IOField "I/O field_108" at 1072,271 size 60x22; FormatPattern 999
   TextField "Text field_58" at 650,271 size 54x22; Text 'IW822'
   TextField "Text field_59" at 703,311 size 220x22; Text 'R3_SPR_AI_824'
   IOField "I/O field_111" at 930,311 size 70x22; FormatPattern 999
      ProcessValue <- "12_AI_Data_R3_SPR_AI_824_SCALED"
   TextField "Text field_60" at 650,311 size 53x22; Text 'IW824'
   TextField "Text field_61" at 703,351 size 220x22; Text 'R3_SPR_AI_826'
   IOField "I/O field_116" at 930,351 size 70x22; FormatPattern 999
      ProcessValue <- "12_AI_Data_R3_SPR_AI_826_SCALED"
   TextField "Text field_62" at 650,351 size 53x22; Text 'IW826'
   TextField "Text field_63" at 703,391 size 220x22; Text 'R3_SPR_AI_828'
   IOField "I/O field_121" at 930,391 size 70x22; FormatPattern 999
      ProcessValue <- "12_AI_Data_R3_SPR_AI_828_SCALED"
   TextField "Text field_64" at 650,391 size 53x22; Text 'IW828'
   TextField "Text field_41" at 133,124 size 89x20; Text 'Description'
   TextField "Text field_42" at 771,124 size 89x20; Text 'Description'
   TextField "Text field_43" at 17,124 size 37x20; Text 'AI'
   TextField "Text field_44" at 661,124 size 37x20; Text 'AI'
   TextField "Text field_47" at 702,431 size 220x22; Text 'R3_SPR_AI_830'
   IOField "I/O field_81" at 929,431 size 70x22; FormatPattern 999
      ProcessValue <- "12_AI_Data_R3_SPR_AI_830_SCALED"
   TextField "Text field_48" at 649,431 size 53x22; Text 'IW830'
   IOField "I/O field_109" at 1140,271 size 60x22; Authorization "Parameter Change"; FormatPattern 999
   IOField "I/O field_110" at 1208,271 size 60x22; Authorization "Parameter Change"; FormatPattern 999
   TextField "Text field_52" at 17,91 size 259x26; Text 'GCU Control PLC (Rack 3)'
   Button "Button_1" at 1160,732 size 100x35; TextOn 'BWTS Digital Inputs.'; TextOff 'Next'
      on Click: ActivateScreen("BC Analogue Inputs", 0)
   TextField "Text field_25" at 60,231 size 220x22; Text 'TIT408 FCW TEMP'
   IOField "I/O field_52" at 361,231 size 60x22; Authorization "Parameter Change"; FormatPattern 999
   IOField "I/O field_53" at 429,231 size 60x22; Authorization "Parameter Change"; FormatPattern 999
   IOField "I/O field_54" at 497,231 size 60x22; Authorization "Parameter Change"; FormatPattern 999
      ProcessValue <- "84_Setpoints_TIT408_High"
   IOField "I/O field_55" at 565,231 size 60x22; Authorization "Parameter Change"; FormatPattern 999
      ProcessValue <- "84_Setpoints_TIT408_HighHigh"
   TextField "Text field_33" at 60,391 size 220x22; Text 'PIT358 FCW INLET PRESS'
   IOField "I/O field_57" at 361,391 size 60x22; Authorization "Parameter Change"; FormatPattern 99.9
      ProcessValue <- "19_AUTO_CMNDS_Data_PIT358_CMND_LowLow"
   IOField "I/O field_58" at 429,391 size 60x22; Authorization "Parameter Change"; FormatPattern 99.9
      ProcessValue <- "19_AUTO_CMNDS_Data_PIT358_CMND_Low"
   IOField "I/O field_59" at 497,391 size 60x22; Authorization "Parameter Change"; FormatPattern 99.9
      ProcessValue <- "19_AUTO_CMNDS_Data_PIT358_CMND_High"
   IOField "I/O field_60" at 565,391 size 60x22; Authorization "Parameter Change"; FormatPattern 99.9
      ProcessValue <- "19_AUTO_CMNDS_Data_PIT358_CMND_HighHigh"
   IOField "I/O field_47" at 1004,191 size 60x22; Authorization "Commissioning"; FormatPattern 9.9
   IOField "I/O field_48" at 1072,191 size 60x22; Authorization "Commissioning"; FormatPattern 9.9
   TextField "Text field_35" at 61,191 size 220x22; Text 'R3_SPR_AI_802'
   IOField "I/O field_49" at 1004,231 size 60x22; FormatPattern 999
   IOField "I/O field_51" at 1072,231 size 60x22; FormatPattern 999
   IOField "I/O field_66" at 1140,231 size 60x22; FormatPattern 999
      ProcessValue <- "84_Setpoints_E400_TT002_High"
   IOField "I/O field_67" at 1208,231 size 60x22; FormatPattern 999
      ProcessValue <- "84_Setpoints_E400_TT002_HighHigh"
   TextField "Text field_37" at 61,349 size 220x22; Text 'PIT416 GAS TO DECK PRESS'
   IOField "I/O field_69" at 362,349 size 60x22; Authorization "Parameter Change"; FormatPattern 9.9
      ProcessValue <- "84_Setpoints_PIT416_LowLow"
   IOField "I/O field_70" at 430,349 size 60x22; Authorization "Parameter Change"; FormatPattern 9.9
      ProcessValue <- "84_Setpoints_PIT416_Low"
   IOField "I/O field_71" at 498,349 size 60x22; Authorization "Parameter Change"; FormatPattern 9.9
      ProcessValue <- "84_Setpoints_PIT416_High"
   IOField "I/O field_72" at 566,349 size 60x22; Authorization "Parameter Change"; FormatPattern 9.9
      ProcessValue <- "84_Setpoints_PIT416_HighHigh"
   TextField "Text field_39" at 1109,687 size 151x62; Text 'To BC Analogue Inputs'
   IOField "I/O field_21" at 1004,310 size 60x22; FormatPattern 999
   IOField "I/O field_22" at 1072,310 size 60x22; FormatPattern 999
   IOField "I/O field_23" at 1140,310 size 60x22; FormatPattern 999
   IOField "I/O field_24" at 1208,310 size 60x22; FormatPattern 999
   IOField "I/O field_25" at 1004,351 size 60x22; FormatPattern 999
   IOField "I/O field_26" at 1072,351 size 60x22; FormatPattern 999
   IOField "I/O field_27" at 1140,351 size 60x22; FormatPattern 999
   IOField "I/O field_28" at 1208,351 size 60x22; FormatPattern 999
   IOField "I/O field_29" at 1004,391 size 60x22; FormatPattern 999
   IOField "I/O field_30" at 1072,391 size 60x22; FormatPattern 999
   IOField "I/O field_31" at 1140,391 size 60x22; FormatPattern 999
   IOField "I/O field_32" at 1208,391 size 60x22; FormatPattern 999
   IOField "I/O field_33" at 1004,430 size 60x22; FormatPattern 999
   IOField "I/O field_34" at 1072,430 size 60x22; FormatPattern 999
   IOField "I/O field_35" at 1140,430 size 60x22; FormatPattern 999
   IOField "I/O field_36" at 1208,430 size 60x22; FormatPattern 999
   IOField "I/O field_37" at 286,191 size 70x22; FormatPattern 999
      ProcessValue <- "12_AI_Data_R3_SPR_AI_802_SCALED"
   IOField "I/O field_38" at 361,190 size 60x22; FormatPattern 999
   IOField "I/O field_39" at 429,190 size 60x22; FormatPattern 999
   IOField "I/O field_40" at 497,190 size 60x22; FormatPattern 999
   IOField "I/O field_50" at 565,190 size 60x22; FormatPattern 999
   IOField "I/O field_56" at 287,231 size 70x22; FormatPattern s999; Unit  °C
      ProcessValue <- "12_AI_Data_TIT_408_SCALED"
   IOField "I/O field_63" at 287,391 size 70x22; FormatPattern s99.9; Unit  Barg
      ProcessValue <- "12_AI_Data_PIT_358_SCALED"
   IOField "I/O field_64" at 287,349 size 70x22; FormatPattern s9.9; Unit  Barg
      ProcessValue <- "12_AI_Data_PIT_416_SCALED"
   Button "Button_2" at 361,391 size 264x22; TextOff 'Text'; Authorization "Commissioning"
      on Press: ActivateScreen("GCU Target Setpoints", 0)
   Button "Button_3" at 362,310 size 264x22; TextOff 'Text'; Authorization "Commissioning"
      on Press: ActivateScreen("GCU Target Setpoints", 0)
   Button "Button_4" at 1004,151 size 264x22; TextOff 'Text'; Authorization "Commissioning"
      on Press: ActivateScreen("GCU Target Setpoints", 0)
   Button "Button_5" at 362,148 size 264x28; TextOff 'Text'; Authorization "Commissioning"
      on Press: ActivateScreen("GCU Target Setpoints", 0)
   Group "Group" at 455,41 size 373x50
   Button "HmiScreenItemData_8" at 469,45 size 355x40; TextOn 'Back'; TextOff 'Text'
   TextField "Screen title" at 455,41 size 373x50; Text 'Screen title'

PopupScreen "Salinity - Acceptance" 1050x350
   Button "Button_2" at 556,290 size 105x50; TextOff 'NO'
      on Release: ActivateScreen("Balast Water Treatment Setup", 0)
   Button "Button_3" at 390,290 size 105x50; TextOff 'YES'
      on Press: function_b14e0dd5("80_From_HMI_SAL_CNFRM", 0)
      on Release: function_efd93a16("Salinity - Acceptance", 168, 315, -1, -1, 1)
   TextField "Text field_1" at 223,102 size 604x82; Text 'Please confirm that the entered salinity value of is correct'
   IOField "I/O field_1" at 510,138 size 139x50; FormatPattern 99.9; Unit  psu
      ProcessValue <- "80_From_HMI_SAL_VALUE"

PopupScreen "PGC Commissioning" 1280x800
   Button "Button_1" at 308,285 size 665x230; TextOff 'Text'
      on Release: ActivateScreen("Inert Gas Generator Plant", 0)
   Button "Button_2" at 540,431 size 200x55; TextOff 'OK'
      on Release: ResetBit("PGC_COMMISSION_MODE_DB_Active")
   TextField "Text field_1" at 303,313 size 674x100; Text 'Tanks can now be changed over, press OK when completed'

PopupScreen "Treatment check / Daily Checks Completed" 1050x350
   Button "Button_3" at 411,283 size 229x50; TextOff 'CONFIRM'
      on Release: function_efd93a16("Treatment check / Daily Checks Completed", 0, 0, 0, -1, 1)
      on Press: function_b14e0dd5("88_treatment_POP_UP_CNFRM", 0)
   TextField "Text field_1" at 3,36 size 1044x240; Text 'Please confirm pre treatment check and daily checks are completed.'

